   *)
END_FUNCTION_BLOCK

FUNCTION_BLOCK "DELAY_4"   // FB108, SCL
TITLE = DELAY_4
{ S7_Optimized_Access := 'FALSE' }
AUTHOR : hugo
FAMILY : SIGPRO
NAME : DELAY4
VERSION : 1.1
// this function block delays input values by each programm cycle
// after 4 cycles the in value has shifted to the out 4 and will be discarded after the next cycle
// the blocks can be cascaded.
   VAR_INPUT
      in : Real;
   END_VAR
   VAR_OUTPUT
      out1 : Real;
      out2 : Real;
      out3 : Real;
      out4 : Real;
   END_VAR
   VAR
      temp : Real;
   END_VAR
BEGIN


     #out4 := #out3;
     #out3 := #out2;
     #out2 := #out1;
     #out1 := #temp;
     #temp := #in;

   (* revision history

   hm 19.1.2007    rev 1.1
       added variable temp to add 1 delay  for q1

   *)
END_FUNCTION_BLOCK

FUNCTION_BLOCK "FADE"   // FB109, SCL
TITLE = FADE
{ S7_Optimized_Access := 'FALSE' }
AUTHOR : oscat
FAMILY : SIGPRO
NAME : FADE
VERSION : 1.3
// FADE is used to crossfade between the inputs IN1 and IN2. The fade_over time is specified with TF.
// When F = TRUE then Y = IN2 after the time TF, and when F = FALSE then Y = IN1.
// 
// uses: RMP_W [FB105]
//       _RMP_W [FB94] 
//       T_PLC_MS [FC64]
//       STIME [FB64],IDB_STIME [DB64]
   VAR_INPUT
      IN1 : Real;
      IN2 : Real;
      F : Bool;
      TF : Time;
      rst : Bool;
   END_VAR
   VAR_OUTPUT
      Y : Real;
   END_VAR
   VAR
      rmx : "RMP_W";
   END_VAR
BEGIN


   #rmx(RST := #rst AND NOT #F, SET := #rst AND #F, PT := #TF, UP := #F);
   #Y := (#IN2 - #IN1) / 65535.0 * DINT_TO_REAL(WORD_TO_DINT(#rmx.out)) + #IN1;


   (* code for rev 1.1
   IF rst THEN
       rmx(set := F, rst := NOT F);
   ELSIF F AND (NOT rmx.high) THEN
       rmx(PT := TF, UP := TRUE, e := TRUE, rst := FALSE, set := FALSE);
   ELSIF (NOT F) AND (NOT rmx.low) THEN
       rmx(PT := TF, UP := FALSE, e := TRUE, rst := FALSE, set := FALSE);
   ELSE
       rmx(e := FALSE, rst := FALSE, set := FALSE);
   END_IF;
   Y := (WORD_TO_REAL(rmx.out) * in1 + WORD_TO_REAL(FF - rmx.out) * IN2) / FF;
   *)


   (* revision history
   hm  26. dec 2007    rev 1.0
       original version

   hm  18. oct. 2008   rev 1.1
       improved performance
       changed calls for rmp_w because rmp_w has chaged

   hm  17. dec. 2008   rev 1.2
       function of input f was inverted

   hm  24. jan. 2009   rev 1.3
       delted unused var FF
   *)
END_FUNCTION_BLOCK

FUNCTION_BLOCK "FILTER_DW"   // FB110, SCL
TITLE = FILTER_DW
{ S7_Optimized_Access := 'FALSE' }
AUTHOR : hugo
FAMILY : SIGPRO
NAME : FILTDW
VERSION : 1.1
// FILTER_DW is an low pass filter with a programmable time T used for DWORD format.
// 
// uses: T_PLC_MS [FC64]
//       STIME [FB64],IDB_STIME [DB64]
   VAR_INPUT
      X : DWord;
      T : Time;
   END_VAR
   VAR_OUTPUT
      Y : DWord;
   END_VAR
   VAR
      last : DWord;
      tx : DWord;
      init : Bool;
      Yi : Real;
   END_VAR
   VAR_TEMP
      TOP_SI : Struct
         EV_CLASS : Byte;
         EV_NUM : Byte;
         PRIORITY : Byte;
         NUM : Byte;
         TYP2_3 : Byte;
         TYP1 : Byte;
         ZI1 : Word;
         ZI2_3 : DWord;
      END_STRUCT;
      START_UP_SI : Struct
         EV_CLASS : Byte;
         EV_NUM : Byte;
         PRIORITY : Byte;
         NUM : Byte;
         TYP2_3 : Byte;
         TYP1 : Byte;
         ZI1 : Word;
         ZI2_3 : DWord;
      END_STRUCT;
      ERR : Int;
   END_VAR
BEGIN


   (* read actual startup info *)
   (* OB1_SCAN_1  BYTE  -  B#16#01: Abschluss des Neustarts (Warmstarts)
                        -  B#16#02: Abschluss des Wiederanlaufs
                        -  B#16#03: Abschluss des freien Zyklus
                        -  B#16#04: Abschluss des Kaltstarts
                        -  B#16#05: Erster OB 1-Zyklus der neuen Master-CPU nach 
                                    Master-Reserve-Umschaltung und STOP des 
                                    bisherigen Masters *)

   #ERR := RD_SINFO (TOP_SI => #TOP_SI, START_UP_SI => #START_UP_SI);

   (* read system time *)
   #tx := "T_PLC_MS"();

   (* reset last_time on system startup *)
   IF #TOP_SI.EV_NUM = 1 OR #TOP_SI.EV_NUM = 2 OR #TOP_SI.EV_NUM = 4 THEN 
       #last := #tx;
   END_IF;

   (* startup initialisation *)
   IF NOT #init OR #T = t#0s THEN
       #init := TRUE;
       #Yi := DWORD_TO_REAL(#X);
   ELSE
       #Yi := #Yi + (DWORD_TO_REAL(#X) - DWORD_TO_REAL(#Y)) * DINT_TO_REAL(DWORD_TO_DINT(#tx) - DWORD_TO_DINT(#last)) / DINT_TO_REAL(T_CONV(#T));
   END_IF;
   #last := #tx;

   #Y := REAL_TO_DWORD(#Yi);


   (*
   hm 10. oct. 2008    rev 1.0
       original version

   hm  3. nov. 2008    REV 1.1
       corrected an overflow problem
   *)
END_FUNCTION_BLOCK

FUNCTION_BLOCK "FILTER_MAV_DW"   // FB111, SCL
TITLE = FILTER_MAV_DW
{ S7_Optimized_Access := 'FALSE' }
AUTHOR : hugo
FAMILY : SIGPRO
NAME : FIMAVDW
VERSION : 1.3
// FILTER_MAV_DW is a moving average filter with programmable length N for DWORD Data.
//  
// uses: INC1 [FC53]
   VAR_INPUT
      X : DWord;
      N : Int;
      RST : Bool;
   END_VAR
   VAR_OUTPUT
      Y : DWord;
   END_VAR
   VAR
      init : Bool;
      buffer : Array[0..31] of DWord;
      i : Int;
   END_VAR
   VAR_TEMP
      tmp : Int;
      tN : Int;
   END_VAR
BEGIN


   (* limit N to size of buffer *)
   #tN := MIN(IN1:=#N, IN2:=32);

   (* startup initialisation *)
   IF NOT #init OR #RST OR #tN = 0 THEN
       #init := TRUE;
       #tmp := #tN - 1;
       FOR #i := 0 TO #tmp DO
           #buffer[#i] := #X;
       END_FOR;
       #Y := #X;
   ELSE
       #tmp := #tN;
       #i := "INC1"(X:=#i, N:=#tmp);
       #Y := DINT_TO_DWORD(DWORD_TO_DINT(#Y) + (DWORD_TO_DINT(#X) - DWORD_TO_DINT(#buffer[#i])) / INT_TO_DINT(#tN));
       #buffer[#i] := #X;
   END_IF;


   (*
   hm 13. oct. 2008    rev 1.0
       original version

   hm  27. oct. 2008   rev 1.1
       added typecast to avoid warnings

   hm  24. nov. 2008   rev 1.2
       added typecasts to avoid warnings
       avoid divide by 0 if N = 0

   hm  23. feb. 2009   rev 1.3
       limit N to max array size

   *)
END_FUNCTION_BLOCK

FUNCTION_BLOCK "FILTER_MAV_W"   // FB112, SCL
TITLE = FILTER_MAV_W
{ S7_Optimized_Access := 'FALSE' }
AUTHOR : hugo
FAMILY : SIGPRO
NAME : FIMAVW
VERSION : 1.4
// FILTER_MAV_W is a moving average filter with programmable length N for WORD Data.
//  
// uses: INC1 [FC53]
   VAR_INPUT
      X : Word;
      N : Int;
      RST : Bool;
   END_VAR
   VAR_OUTPUT
      Y : Word;
   END_VAR
   VAR
      init : Bool;
      buffer : Array[0..31] of Word;
      i : Int;
      sum : DWord;
   END_VAR
   VAR_TEMP
      tmp : Int;
      tN : Int;
   END_VAR
BEGIN


   (* limit N to size of buffer *)
   #tN := MIN(IN1:=#N, IN2:=32);

   (* startup initialisation *)
   IF NOT #init OR #RST OR #tN = 0 THEN
     #init := TRUE;
     #tmp := #tN - 1;
     FOR #i := 0 TO #tmp DO
       #buffer[#i] := #X;
     END_FOR;
     #sum := DINT_TO_DWORD(WORD_TO_DINT(#Y) * INT_TO_DINT(#tN));
     #Y := #X;
   ELSE
     #tmp := #tN;
     #i := "INC1"(X:=#i, N:=#tmp);
     #sum := DINT_TO_DWORD(DWORD_TO_DINT(#sum) + WORD_TO_DINT(#X) - WORD_TO_DINT(#buffer[#i]));
     #Y := DINT_TO_WORD(DWORD_TO_DINT(#sum) / INT_TO_DINT(#tN));
     #buffer[#i] := #X;
   END_IF;


   (*
   hm 13. oct. 2008  rev 1.0
     original version

   hm  18. oct. 2008 rev 1.1
     added typecast to avoid warnings

   hm  24. nov. 2008 rev 1.2
     added typecasts to avoid warnings
     avoid devide by 0 if N = 0

   hm  23. feb. 2009 rev 1.3
     limit N to max array size

   hm  26. mar. 2011 rev 1.4
     corrected error in calculation
   *)
END_FUNCTION_BLOCK

FUNCTION_BLOCK "FILTER_W"   // FB113, SCL
TITLE = FILTER_W
{ S7_Optimized_Access := 'FALSE' }
AUTHOR : hugo
FAMILY : SIGPRO
NAME : FILTW
VERSION : 1.2
// FILTER_DW is an low pass filter with a programmable time T used for DWORD format.
// 
// uses: T_PLC_MS [FC64]
//       STIME [FB64],IDB_STIME [DB64]
   VAR_INPUT
      X : Word;
      T : Time;
   END_VAR
   VAR_OUTPUT
      Y : Word;
   END_VAR
   VAR
      last : DWord;
      tx : DWord;
      init : Bool;
      tmp : DWord;
   END_VAR
   VAR_TEMP
      TOP_SI : Struct
         EV_CLASS : Byte;
         EV_NUM : Byte;
         PRIORITY : Byte;
         NUM : Byte;
         TYP2_3 : Byte;
         TYP1 : Byte;
         ZI1 : Word;
         ZI2_3 : DWord;
      END_STRUCT;
      START_UP_SI : Struct
         EV_CLASS : Byte;
         EV_NUM : Byte;
         PRIORITY : Byte;
         NUM : Byte;
         TYP2_3 : Byte;
         TYP1 : Byte;
         ZI1 : Word;
         ZI2_3 : DWord;
      END_STRUCT;
      ERR : Int;
   END_VAR
BEGIN


   (* read actual startup info *)
   (* OB1_SCAN_1  BYTE  -  B#16#01: Abschluss des Neustarts (Warmstarts)
                        -  B#16#02: Abschluss des Wiederanlaufs
                        -  B#16#03: Abschluss des freien Zyklus
                        -  B#16#04: Abschluss des Kaltstarts
                        -  B#16#05: Erster OB 1-Zyklus der neuen Master-CPU nach 
                                    Master-Reserve-Umschaltung und STOP des 
                                    bisherigen Masters *)

   #ERR := RD_SINFO (TOP_SI => #TOP_SI, START_UP_SI => #START_UP_SI);

   (* read system time *)
   #tx := "T_PLC_MS"();

   (* reset last_time on system startup *)
   IF #TOP_SI.EV_NUM = 1 OR #TOP_SI.EV_NUM = 2 OR #TOP_SI.EV_NUM = 4 THEN 
     #init := false;
   END_IF;

   (* startup initialisation *)
   IF NOT #init OR #T = t#0s THEN
     #init := TRUE;
     #last := #tx;
     #Y := #X;
   ELSIF #Y = #X THEN
     #last := #tx;
   ELSE
     #tmp :=  DINT_TO_DWORD((WORD_TO_DINT(#X) - WORD_TO_DINT(#Y)) * (DWORD_TO_DINT(#tx) - DWORD_TO_DINT(#last)) / T_CONV(#T));
     IF #tmp <> 0 THEN
       #Y := DINT_TO_WORD(WORD_TO_DINT(#Y) + DWORD_TO_DINT(#tmp));
       #last := #tx;
     END_IF;
   END_IF;


   (*
   hm 10. oct. 2008  rev 1.0
     original version

   hm  3. nov. 2008  rev 1.1
     fixed overflow problem in formula

   hm  25. jan. 2011 rev 1.2
     fixed error in formula
   *)
END_FUNCTION_BLOCK

FUNCTION_BLOCK "FILTER_WAV"   // FB114, SCL
TITLE = FILTER_WAV
{ S7_Optimized_Access := 'FALSE' }
AUTHOR : hugo
FAMILY : SIGPRO
NAME : FILTWAV
VERSION : 1.2
// FILTER_WAV is a moving average filter with programmable length N for DWORD Data.
// 
// uses: INC1 [FC53]
//       DEC1 [FC52]
   VAR_INPUT
      X : Real;
      W : Array[0..15] of Real;
      RST : Bool;
   END_VAR
   VAR_OUTPUT
      Y : Real;
   END_VAR
   VAR
      init : Bool;
      buffer : Array[0..15] of Real;
      i : Int;
      n : Int;
   END_VAR
BEGIN


   (* startup initialisation *)
   IF NOT #init OR #RST THEN
       #init := TRUE;
       FOR #i := 0 TO 15 DO
           #buffer[#i] := #X;
       END_FOR;
       #i := 15;
       #Y := #X;
   ELSE
       #i := "INC1"(N:=16, X:=#i);
       #buffer[#i] := #X;
   END_IF;

   (* calculate the weighted average *)
   #Y := 0.0;
   FOR #n := 0 TO 15 DO
       #Y := #buffer[#i] * #W[#n] + #Y;
       #i := "DEC1"(N:=16, X:=#i);
   END_FOR;


   (*
   hm  14. oct. 2008   rev 1.0
       original version

   hm  27. oct. 2008   rev 1.1
       changed _DEC and _INC to DEC1 and INC1

   hm  10. mar. 2009   rev 1.2
       real constants updated to new systax using dot

   *)
END_FUNCTION_BLOCK

FUNCTION_BLOCK "SEL2_OF_3"   // FB115, SCL
TITLE = SEL2_OF_3
{ S7_Optimized_Access := 'FALSE' }
AUTHOR : oscat
FAMILY : SIGPRO
NAME : SEL2OF3
VERSION : 1.1
// SEL2_OF_3 checks if 3 input Signals are within a distance D from each other and calculates the average of the 3 inputs do not offset more than D from each other.
// If 1 input is more than D greater or smaller than any other input it will be ignored and the average will be calcualted from the remaining 2 Inputs.
// In the case the Output is only calculated from 2 Inputs a Warning Output W will display the Number of the discarded Input. if none of the 3 Inputs are within the allowed Delata D from each other, 
// an Error Output E is set True and the last valid Output will remain active until at least 2 Inputs are within a valid Range from each other.
   VAR_INPUT
      IN1 : Real;
      IN2 : Real;
      IN3 : Real;
      D : Real;
   END_VAR
   VAR_OUTPUT
      Y : Real;
      W : Int;
      "E" : Bool;
   END_VAR
   VAR
      D12 : Bool;
      D23 : Bool;
      D31 : Bool;
   END_VAR
BEGIN


   #D12 := ABS(#IN1-#IN2) <= #D;
   #D23 := ABS(#IN2-#IN3) <= #D;
   #D31 := ABS(#IN3-#IN1) <= #D;

   IF (#D12 AND #D23) OR (#D12 AND #D31) OR (#D23 AND #D31) THEN
       (* all 3 inputs are valid *)
       #Y := (#IN1 + #IN2 + #IN3) * 0.333333333333;
       #"E" := FALSE;
       #W := 0;
   ELSIF #D12 THEN
       (* only inut 1 and 2 are valid *)
       #Y := (#IN1 + #IN2) * 0.5;
       #"E" := FALSE;
       #W := 3;
   ELSIF #D23 THEN
       (* only inut 2 and 3 are valid *)
       #Y := (#IN2 + #IN3) * 0.5;
       #"E" := FALSE;
       #W := 1;
   ELSIF #D31 THEN
       (* only inut 3 and 1 are valid *)
       #Y := (#IN3 + #IN1) * 0.5;
       #"E" := FALSE;
       #W := 2;
   ELSE
       (* no calculation possible *)
       #"E" := TRUE;
       #W := 4;
   END_IF;


   (* revision history
   hm  18. may 2008    rev 1.0
       original version

   hm  10. mar. 2009   rev 1.1
       improved code
   *)
END_FUNCTION_BLOCK

FUNCTION_BLOCK "SEL2_OF_3B"   // FB116, SCL
TITLE = SEL2_OF_3B
{ S7_Optimized_Access := 'FALSE' }
AUTHOR : oscat
FAMILY : SIGPRO
NAME : SEL2OF3B
VERSION : 1.0
// SEL2_OF_3B is used to connect 3 binary sensors to one signal. the output Q reflects the state of at least two inputs.
// if two or more of the 3 inputs ate TRUE then Q will be TRUE and if two or more of the three inputs are FALSE then Q will be false.
// the main putrpose is the connection of 3 redundant binary sensors.  
// The output W will be active when one of the 3 inputs is of different state.
// to avoid flickering while the sensors are switching the output W will become active after a programmed delay of TD.
   VAR_INPUT
      IN1 : Bool;
      IN2 : Bool;
      IN3 : Bool;
      TD : Time;
   END_VAR
   VAR_OUTPUT
      Q : Bool;
      W : Bool;
   END_VAR
   VAR
      TDEL : TON;
   END_VAR
BEGIN


   #Q := (#IN1 AND #IN2) OR (#IN1 AND #IN3) OR (#IN2 AND #IN3);
   #TDEL(IN := (#IN1 XOR #IN2) OR (#IN1 XOR #IN3) OR (#IN2 XOR #IN3), PT := #TD);
   #W := #TDEL.Q;


   (* revision history
   hm      19. may 2008    rev 1.0
       original version

   *)
END_FUNCTION_BLOCK

FUNCTION_BLOCK "SH"   // FB117, SCL
TITLE = SH
{ S7_Optimized_Access := 'FALSE' }
AUTHOR : hugo
FAMILY : SIGPRO
NAME : SH
VERSION : 1.1
// this sample and hold module samples an input at the rising edge of clk an stores it in out.
// the out stays stable until the next rising clk edge appears.
// a trigger output as active for one cycle when the output was updated.
   VAR_INPUT
      in : Real;
      CLK : Bool;
   END_VAR
   VAR_OUTPUT
      out : Real;
      trig : Bool;
   END_VAR
   VAR
      edge : Bool;
   END_VAR
BEGIN


     IF #CLK AND NOT #edge THEN
         #out := #in;
         #trig := TRUE;
     ELSE;
         #trig := FALSE;
     END_IF;
     #edge := #CLK;

   (* revision history

   hm 16.1.2007    rev 1.1
       added trig output

   *)
END_FUNCTION_BLOCK

FUNCTION_BLOCK "SH_1"   // FB118, SCL
TITLE = SH_1
{ S7_Optimized_Access := 'FALSE' }
AUTHOR : hugo
FAMILY : SIGPRO
NAME : SH_1
VERSION : 1.2
// this sample and hold module samples an input every PT seconds.
// after a ample is taken the output Trig will be active for one cycle.
// 
// uses: T_PLC_MS [FC64]
//       STIME [FB64],IDB_STIME [DB64]
   VAR_INPUT
      in : Real;
      PT : Time;
   END_VAR
   VAR_OUTPUT
      out : Real;
      Trig : Bool;
   END_VAR
   VAR
      last : Time;
      tx : Time;
   END_VAR
   VAR_TEMP
      TOP_SI : Struct
         EV_CLASS : Byte;
         EV_NUM : Byte;
         PRIORITY : Byte;
         NUM : Byte;
         TYP2_3 : Byte;
         TYP1 : Byte;
         ZI1 : Word;
         ZI2_3 : DWord;
      END_STRUCT;
      START_UP_SI : Struct
         EV_CLASS : Byte;
         EV_NUM : Byte;
         PRIORITY : Byte;
         NUM : Byte;
         TYP2_3 : Byte;
         TYP1 : Byte;
         ZI1 : Word;
         ZI2_3 : DWord;
      END_STRUCT;
      ERR : Int;
   END_VAR
BEGIN


   (* OB1_SCAN_1  BYTE  -  B#16#01: Abschluss des Neustarts (Warmstarts)
                        -  B#16#02: Abschluss des Wiederanlaufs
                        -  B#16#03: Abschluss des freien Zyklus
                        -  B#16#04: Abschluss des Kaltstarts
                        -  B#16#05: Erster OB 1-Zyklus der neuen Master-CPU nach 
                                    Master-Reserve-Umschaltung und STOP des 
                                    bisherigen Masters *)

   #ERR := RD_SINFO (TOP_SI => #TOP_SI, START_UP_SI => #START_UP_SI);

   (* reset last_time on system startup *)
   IF #TOP_SI.EV_NUM = 1 OR #TOP_SI.EV_NUM = 2 OR #TOP_SI.EV_NUM = 4 THEN 
       #last := t#0ms;
   END_IF;

     (* read system time *)
     #tx := T_CONV(DWORD_TO_DINT("T_PLC_MS"()));

     IF #tx - #last >= #PT THEN
       #last := #tx;
       #out := #in;
       #Trig := TRUE;
     ELSE
       #Trig := FALSE;
     END_IF;

   (* revision history

   HM  6.1.2007  rev 1.1
     added trig output

   HM  17.9.2007  rev 1.2
     replaced time() with T_PLC_MS() for compatibility reasons
   *)
END_FUNCTION_BLOCK

FUNCTION_BLOCK "SH_2"   // FB119, SCL
TITLE = SH_2
{ S7_Optimized_Access := 'FALSE' }
AUTHOR : hugo
FAMILY : SIGPRO
NAME : SH_2
VERSION : 1.6
// this sample and hold module samples an input every PT seconds.
// this sample and hold also does avg and other calculations with the input data.
// an average is calculated while for this calculation disc samples are discarded,
// disc = 0 all samples are averaged,
// if disc = 1 the lowest value is ignored,
// if disc = 2 the lowest and highest values are ignored, 
// and so on.....
// 
// uses: T_PLC_MS [FC64]
//       STIME [FB64],IDB_STIME [DB64]
//       EVEN [FC76]
   VAR_INPUT
      in : Real;
      PT : Time;
      N : Int := 16;
      disc : Int;
   END_VAR
   VAR_OUTPUT
      out : Real;
      trig : Bool;
      avg : Real;
      high : Real;
      low : Real;
   END_VAR
   VAR
      "M" : Int;
      buf : Array[0..15] of Real;
      buf2 : Array[0..15] of Real;
      last : Time;
      i : Int;
      start : Int;
      temp : Real;
      stop : Int;
      tx : Time;
      d2 : Int;
   END_VAR
   VAR_TEMP
      TOP_SI : Struct
         EV_CLASS : Byte;
         EV_NUM : Byte;
         PRIORITY : Byte;
         NUM : Byte;
         TYP2_3 : Byte;
         TYP1 : Byte;
         ZI1 : Word;
         ZI2_3 : DWord;
      END_STRUCT;
      START_UP_SI : Struct
         EV_CLASS : Byte;
         EV_NUM : Byte;
         PRIORITY : Byte;
         NUM : Byte;
         TYP2_3 : Byte;
         TYP1 : Byte;
         ZI1 : Word;
         ZI2_3 : DWord;
      END_STRUCT;
      ERR : Int;
   END_VAR
BEGIN


   (* read actual startup info *)
   (* OB1_SCAN_1  BYTE  -  B#16#01: Abschluss des Neustarts (Warmstarts)
                        -  B#16#02: Abschluss des Wiederanlaufs
                        -  B#16#03: Abschluss des freien Zyklus
                        -  B#16#04: Abschluss des Kaltstarts
                        -  B#16#05: Erster OB 1-Zyklus der neuen Master-CPU nach 
                                    Master-Reserve-Umschaltung und STOP des 
                                    bisherigen Masters *)

   #ERR := RD_SINFO (TOP_SI => #TOP_SI, START_UP_SI => #START_UP_SI);

   (* reset last_time on system startup *)
   IF #TOP_SI.EV_NUM = 1 OR #TOP_SI.EV_NUM = 2 OR #TOP_SI.EV_NUM = 4 THEN 
       #last := t#0ms;
   END_IF;

   (* read system time *)
   #tx := T_CONV(DWORD_TO_DINT("T_PLC_MS"()));
   #d2 := WORD_TO_INT(SHR(IN:=INT_TO_WORD(#disc),N:=1));

   IF #tx - #last >= #PT THEN
       #last := #tx;
       #trig := TRUE;

       (* limit M to 0..16 *)
       #"M" := LIMIT(MN:=1,IN:=#N,MX:=16);

       (* edge detected lets take the sample *)
       FOR #i := #"M" - 1 TO 1 BY -1 DO #buf2[#i] := #buf2[#i-1]; END_FOR;
       #buf2[0] := #in;
       #out := #in;
       #buf BLKMOV #buf2;

       (* sort the ARRAY lowest value AT 0 *)
       FOR #start := 0 TO #"M" - 2 DO
         FOR #i := #start+1 TO #"M" - 1 DO
           IF #buf[#start] > #buf[#i] THEN
             #temp := #buf[#start];
             #buf[#start] := #buf[#i];
             #buf[#i] := #temp;
           END_IF;
         END_FOR;
       END_FOR;

       (* any calculation with the samples is here *)
       #stop := #"M" - 1 - #d2;
       #start := #d2;
       IF NOT "EVEN"(#disc) THEN #start := #start + 1; END_IF;
       #avg := 0;
       FOR #i := #start TO #stop DO #avg := #avg + #buf[#i]; END_FOR;
       #avg := #avg / INT_TO_REAL(#stop - #start +1);
       #low := #buf[#start];
       #high := #buf[#stop];
   ELSE
       #trig := FALSE;
   END_IF;


   (* revision history
   hm 20. jan. 2007    rev 1.1
       added input N to specify the amout of samples for average and high low calculations
       added trig output

   hm 10. sep. 2007    rev 1.2
       an error would be generated if N was set to 0, now n is forced to1 if set to 0.
       index was out of array.

   hm  17. sep. 2007   rev 1.3
       replaced time() with t_plc_ms() for compatibility reasons

   hm  6. jan. 2008    rev 1.4
       improved performance

   hm  14. jun. 2008   rev 1.5
       set default for input N = 16

   hm  10. mar. 2009   rev 1.6
       added type conversion for compatibility reasons

   *)
END_FUNCTION_BLOCK

FUNCTION_BLOCK "SH_T"   // FB120, SCL
TITLE = SH_T
{ S7_Optimized_Access := 'FALSE' }
AUTHOR : hugo
FAMILY : SIGPRO
NAME : SH_T
VERSION : 1.1
// this sample and hold module samples an input while en is high.
// during the high time of en the output follows in.
// the out stays stable until the en goes high again.
   VAR_INPUT
      IN : Real;
      "E" : Bool;
   END_VAR
   VAR_OUTPUT
      OUT : Real;
   END_VAR
BEGIN


   IF #"E" THEN #OUT := #IN; END_IF;

   (* revision history
   hm  1. sep. 2006    rev 1.0
       original version

   hm  18. oct. 2008   rev 1.1
       changed input en to e for compatibility reasons

   *)
END_FUNCTION_BLOCK

FUNCTION_BLOCK "STAIR2"   // FB121, SCL
TITLE = STAIR2
{ S7_Optimized_Access := 'FALSE' }
AUTHOR : oscat
FAMILY : SIGPRO
NAME : STAIR2
VERSION : 1.4
// the function stair2 converts an anlog input signal to a staircase like output.
// D is the step width for the output signal. the output will use D as a hysteresis for a stairchange.
// if D = 0 then the output follows the input without a chage.
// 
// uses: FLOOR [FC81]
   VAR_INPUT
      X : Real;
      D : Real;
   END_VAR
   VAR_OUTPUT
      Y : Real;
   END_VAR
BEGIN


   IF #D > 0.0 THEN
       IF #X >= #Y + #D OR #X <= #Y - #D THEN #Y := "FLOOR"(#X/#D) * #D; END_IF;
   ELSE
       #Y := #X;
   END_IF;


   (* revision history
   hm  28 jan 2007     rev 1.0
       original version

   hm  27. dec 2007    rev 1.1
       changed code for better performance

   hm  30. jun. 2008   rev 1.2
       added type conversions to avoid warnings under codesys 3.0

   ks  26. oct. 2008   rev 1.3
       improved code

   hm  10. mar. 2009   rev 1.4
       real constants updated to new systax using dot

   *)
END_FUNCTION_BLOCK

FUNCTION_BLOCK "FILTER_I"   // FB238, SCL
TITLE = FILTER_I
{ S7_Optimized_Access := 'FALSE' }
AUTHOR : hugo
FAMILY : SIGPRO
NAME : FILTI
VERSION : 1.0
// FILTER_I is a low pass filter with a programmable time T used for INT format.
//  
// uses: T_PLC_MS [FC64]
//       STIME [FB64],IDB_STIME [DB64]
   VAR_INPUT
      X : Int;
      T : Time;
   END_VAR
   VAR_OUTPUT
      Y : Int;
   END_VAR
   VAR
      Yi : DInt;
      last : DWord;
      tx : DWord;
      init : Bool;
   END_VAR
   VAR_TEMP
      TOP_SI : Struct
         EV_CLASS : Byte;
         EV_NUM : Byte;
         PRIORITY : Byte;
         NUM : Byte;
         TYP2_3 : Byte;
         TYP1 : Byte;
         ZI1 : Word;
         ZI2_3 : DWord;
      END_STRUCT;
      START_UP_SI : Struct
         EV_CLASS : Byte;
         EV_NUM : Byte;
         PRIORITY : Byte;
         NUM : Byte;
         TYP2_3 : Byte;
         TYP1 : Byte;
         ZI1 : Word;
         ZI2_3 : DWord;
      END_STRUCT;
      ERR : Int;
   END_VAR
BEGIN


   (* read actual startup info *)
   (* OB1_SCAN_1  BYTE  -  B#16#01: Abschluss des Neustarts (Warmstarts)
                        -  B#16#02: Abschluss des Wiederanlaufs
                        -  B#16#03: Abschluss des freien Zyklus
                        -  B#16#04: Abschluss des Kaltstarts
                        -  B#16#05: Erster OB 1-Zyklus der neuen Master-CPU nach 
                                    Master-Reserve-Umschaltung und STOP des 
                                    bisherigen Masters *)

   #ERR := RD_SINFO (TOP_SI => #TOP_SI, START_UP_SI => #START_UP_SI);

   (* read system time *)
   #tx := "T_PLC_MS"();

   (* reset last_time on system startup *)
   IF #TOP_SI.EV_NUM = 1 OR #TOP_SI.EV_NUM = 2 OR #TOP_SI.EV_NUM = 4 THEN 
       #last := #tx;
   END_IF;

   (* startup initialisation *)
   IF NOT #init OR #T = t#0s THEN
       #init := TRUE;
       #Yi := INT_TO_DINT(#X) * 1000;
   ELSE
       (* to increase accuracy of the filter we calculate internal Yi wich is Y * 1000 *)
       #Yi := #Yi + INT_TO_DINT(#X - #Y) * (DWORD_TO_DINT(#tx) - DWORD_TO_DINT(#last)) * 1000 / T_CONV(#T);
   END_IF;
   #last := #tx;
   #Y := DINT_TO_INT(#Yi / 1000);


   (*
   hm 8. nov. 2008 rev 1.0
       original version

   *)
END_FUNCTION_BLOCK

FUNCTION_BLOCK "TREND_DW"   // FB245, SCL
TITLE = TREND_DW
{ S7_Optimized_Access := 'FALSE' }
AUTHOR : hugo
FAMILY : SIGPRO
NAME : TREND_DW
VERSION : 1.2
// trend_DW analyses the trend of a input signal.
// The Output Q is True if the input X is >= last_X and is false if the input X is <= last_X
// in addition to the trend the output TU will be high for one cycle to signal a rising of the input value X
// and  TD will signal a decreasing value on the input X.
// in case of a change the output D will show the delta of the input to the last input value.
   VAR_INPUT
      X : DWord;
   END_VAR
   VAR_OUTPUT
      Q : Bool;
      TU : Bool;
      TD : Bool;
      D : DWord;
   END_VAR
   VAR
      last_X : DWord;
   END_VAR
BEGIN


   IF DWORD_TO_DINT(#X) > DWORD_TO_DINT(#last_X) THEN
       #TU := TRUE;
       #TD := FALSE;
       #D := DINT_TO_DWORD(DWORD_TO_DINT(#X) - DWORD_TO_DINT(#last_X));
       #Q := TRUE;
   ELSIF DWORD_TO_DINT(#X) < DWORD_TO_DINT(#last_X) THEN
       #TD := TRUE;
       #TU := FALSE;
       #D := DINT_TO_DWORD(DWORD_TO_DINT(#last_X) - DWORD_TO_DINT(#X));
       #Q := FALSE;
   ELSE
       #TU := FALSE; 
       #TD := FALSE;
       #D := 0;
   END_IF;
   #last_X := #X;


   (* revision history
   hm  21. nov. 2008   rev 1.0
       original version

   hm  20. feb. 2009   rev 1.1
       added outputs TU, TD and D

   hm  14. mar. 2009   rev 1.2
       removed double assignments

   *)
END_FUNCTION_BLOCK

FUNCTION_BLOCK "TREND"   // FB251, SCL
TITLE = TREND
{ S7_Optimized_Access := 'FALSE' }
AUTHOR : hugo
FAMILY : SIGPRO
NAME : TREND
VERSION : 1.0
// trend analyses the trend of a input signal.
// The Output Q is True if the input X is >= last_X and is false if the input X is <= last_X
// in addition to the trend the output TU will be high for one cycle to signal a rising of the input value X
// and  TD will signal a decreasing value on the input X.
// in case of a change the output D will show the delta of the input to the last input value.
   VAR_INPUT
      X : Real;
   END_VAR
   VAR_OUTPUT
      Q : Bool;
      TU : Bool;
      TD : Bool;
      D : Real;
   END_VAR
   VAR
      last_X : Real;
   END_VAR
BEGIN


   #TU := #X > #last_X;
   #TD := #X < #last_X;
   #Q := #TU OR #TD;
   #D := #X - #last_X;

   #last_X := #X;



   (* revision history
   hm 21. aug. 2009 rev 1.0
    original version

   *)
END_FUNCTION_BLOCK

FUNCTION "DEC1" : Int   // FC52, SCL
TITLE = DEC1
{ S7_Optimized_Access := 'FALSE' }
AUTHOR : hugo
FAMILY : MATH
NAME : DEC1
VERSION : 1.1
// This is a decrement function which decrements the variable X by 1 and if 0 is reached, it begins with M again.
// _dec1(3,X) will generate 3,2,1,0,3,2,...
   VAR_INPUT
      X : Int;
      N : Int;
   END_VAR
BEGIN


   IF #X = 0 THEN
       #DEC1 := #N - 1;
   ELSE
       #DEC1 := #X - 1;
   END_IF;

   (* this is a very elegant version but 50% slower
   X := (X - 1 + N) MOD N;
   *)


   (* revision history
   hm  13. oct. 2008   rev 1.0
       original version

   hm  27. oct. 2008   rev 1.1
       added statement to return value for compatibility reasons
   *)
END_FUNCTION

FUNCTION "INC1" : Int   // FC53, SCL
TITLE = INC1
{ S7_Optimized_Access := 'FALSE' }
AUTHOR : hugo
FAMILY : MATH
NAME : INC1
VERSION : 1.2
// This is a increment function which increments the variable X by 1 and if M is reached, it begins with 0 again.
// _inc1(3,X) will generate 0,1,2,3,0,1,.....
   VAR_INPUT
      X : Int;
      N : Int;
   END_VAR
BEGIN


   IF #X >= #N - 1 THEN
       #INC1 := 0;
   ELSE
       #INC1 := #X + 1;
   END_IF;


   (* this elegant version is 50% slower
   INC1 := X := (x + 1) MOD N;
   *)



   (* revision history
   hm  13. oct. 2008   rev 1.0
       original version

   hm  22. oct. 2008   rev 1.1
       added statement to return value for compatibility reasons

   hm  23. feb. 2009   rev 1.2
       when inc1 is called with X >= N inc will continue with 0
   *)
END_FUNCTION

FUNCTION "T_PLC_MS" : DWord   // FC64, SCL
TITLE = T_PLC_MS
{ S7_Optimized_Access := 'FALSE' }
AUTHOR : hugo
FAMILY : MEASURE
NAME : T_PLC_MS
VERSION : 1.2
// T_PLC_MS reads the internal PLC timer and return the time, it has the advantage to be able to set a debug mode 
// and speed up the counter to test the plc timer overrun which occurs every 50 days respectively 25 days at siemens S7
// this routine also allows to correct the behavior of s7 where the internal plc counter will not count all 32 bits.
// 
// uses: STIME [FB64],IDB_STIME [DB64]
BEGIN


   "IDB_STIME"(); 
   #T_PLC_MS := "IDB_STIME".tx; 
   (* hier muss die korrektur für step7 stattfinden
   plctime muss den vollen wertebereich von time ausnutzen:
   wenn bei step7 time -24tage bis plus 24 tage ist dann muss der timer auch beim überlauf auf -24tage springen 
   und auf keinen fall auf 0 !!!!
   für siemens muss ein weiterer fb im main eingebunden werden der sicherstellt das alle 32 bits durchgezählt werden.
   es kann nur ein fb sein den er muss sich das oberste (32te) bit merken.
   oder etwa spring s7 bei überlauf auf -24 tage????? dann wäre keine korrektur nötig.
   *)
   IF "debug" THEN
       #T_PLC_MS := DINT_TO_DWORD((DWORD_TO_DINT(SHL(IN:=#T_PLC_MS,N:="N") OR SHL(IN:=DWORD#1,N:="N"))-1) + DWORD_TO_DINT("offset_FC64_1"));
   END_IF;


   (* revision history
   hm  14.9.2007   rev 1.0
       original version

   hm  12. nov 2007    rev 1.1
       added temporaray variable tx because some compilers could not handle time() as an argument

   hm  16. nov. 2008   rev 1.2
       initialized constants with 0 for compatibility reasons
   *)
END_FUNCTION

FUNCTION "EVEN" : Bool   // FC76, SCL
TITLE = EVEN
{ S7_Optimized_Access := 'FALSE' }
AUTHOR : hugo
FAMILY : MATH
NAME : EVEN
VERSION : 1.2
// this function chacks an input for even value
// the output is true if the input is even.
   VAR_INPUT
      in : DInt;
   END_VAR
   VAR_TEMP
      tIN : DInt;
      _IN AT tIN : Array[0..31] of Bool;
   END_VAR
BEGIN


   #tIN := #in;
   #EVEN := NOT #_IN[24]; //EVEN := NOT in.0;

   (* revision history
   hm  1. oct 2006 rev 1.0
     ORIGINAL VERSION

   hm  01.12.2007  rev 1.1
     changed code for improved performance

   hm  21. mar. 2008 rev 1.2
     changed type of input IN from INT to DINT
   *)
END_FUNCTION

FUNCTION "FLOOR" : Int   // FC81, SCL
TITLE = FLOOR
{ S7_Optimized_Access := 'FALSE' }
AUTHOR : hugo
FAMILY : MATH
NAME : FLOOR
VERSION : 1.1
// This is a rounding function which returns the biggest possible integer which is less or equal to X.
// floor(3.14) = 3
// floor(-3.14) = 4
   VAR_INPUT
      X : Real;
   END_VAR
BEGIN


   #FLOOR := REAL_TO_INT(#X);
   IF #FLOOR > #X THEN
       #FLOOR := #FLOOR - 1;
   END_IF;

   (* revision history
   hm    7. feb 2007   rev 1.0
     originlal version

   hm    21. mar. 2008 rev 1.1
     replaced trunc with real_to_int for compatibility reasons

   *)
END_FUNCTION

FUNCTION "SIGN_R" : Bool   // FC109, SCL
TITLE = SIGN_R
{ S7_Optimized_Access := 'FALSE' }
AUTHOR : hugo
FAMILY : MATH
NAME : SIGN_R
VERSION : 1.4
// this function return true if the real input is negative
   VAR_INPUT
      in : Real;
   END_VAR
BEGIN


   #SIGN_R := #in < 0.0;


   (* revision history
   hm 19.1.2007    rev 1.1
       changed method of function for better compatibility to other systems

   hm  1.12.2007   rev 1.2
       changed code to improve performance

   hm  14. jun. 2008   rev 1.3
       improved performace

   hm 10. mar. 2009    rev 1.4
       real constants updated to new systax using dot
   *)
END_FUNCTION

FUNCTION "AIN" : Real   // FC317, SCL
TITLE = AIN
{ S7_Optimized_Access := 'FALSE' }
AUTHOR : oscat
FAMILY : SIGPRO
NAME : AIN
VERSION : 1.5
// Ain converts signals from A/D converters or other analog sources to an internal real value
// the lowest number of bits are extracted from the input word and the sign will be extracted if available separately.
// the output signal is then conditioned to range from low to high values for a 0 to max value on the analog inputs:
// for example a 15bit input (bits := 12) with sign at bit 15 (0..15) will deliver 0.0 (low value at 0) for an input value of 2#0000_0000_0000
// an input value of 2#1111_1111_1111 will deliver 10.0 on the output (high value set to 10).
   VAR_INPUT
      in : DWord;
      Bits : Byte;
      sign : Byte;
      low : Real;
      high : Real;
   END_VAR
   VAR_TEMP
      temp1 : DWord;
      ttemp1 AT temp1 : Array[0..31] of Bool;
      temp2 : DWord;
      sx : Bool;
   END_VAR
BEGIN


     (* extract the sign bit *)
     IF BYTE_TO_INT(#sign) < 32 THEN
         #temp1 := SHR(IN:=#in,N:=BYTE_TO_INT(#sign));
         #sx := #ttemp1[24];
     ELSE
         #sx := FALSE;
     END_IF;
     #temp1 := SHR(IN:="ff",N:=32-BYTE_TO_INT(#Bits));
     #temp2 := #in AND #temp1;
     #AIN := (#high - #low) * DWORD_TO_REAL(#temp2) / DWORD_TO_REAL(#temp1) + #low;
     IF #sx THEN #AIN := -#AIN; END_IF;

   (* revision history
   hm 18.8.2006    rev 1.1
       fixed an error with low value negative and high value 0.

   hm 19.1.2007    rev 1.2
       fixed an error with sign bit.

   hm  13.9.2007   rev 1.3
       changed code to avoid warning under codesys 2.8.1

   hm  2. dec 2007 rev 1.4
       changed code for better performance

   hm  16. mar 2008    rev 1.5
       added type conversions to avoid warnings under codesys 30
   *)
END_FUNCTION

FUNCTION "AOUT" : DWord   // FC318, SCL
TITLE = AOUT
{ S7_Optimized_Access := 'FALSE' }
AUTHOR : oscat
FAMILY : SIGPRO
NAME : AOUT
VERSION : 1.4
// this module conditions an internal real value for a signal output D/A converter.
// Aout converts and internal real value to a word for an D/A converter or other output devices.
// The input value is converted to a n-bit wide output and a sign bit is set separately as specified.
// the outout min value is set for the specified min input value and the max output is set for the max input value.
// an input higher or lower then the max or min value will set the respective max or min value or the output.
// 
// uses: SIGN_R [FC109]
   VAR_INPUT
      in : Real;
      Bits : Byte;
      sign : Byte;
      low : Real;
      high : Real;
   END_VAR
   VAR_TEMP
      in2 : Real;
      sx : Bool;
   END_VAR
BEGIN


     (* if sign bit is defined *)
     IF WORD_TO_INT(BYTE_TO_WORD(#sign)) < 32 THEN
         #sx := "SIGN_R"(in:=#in);
         #in2 := ABS(#in);
     ELSE
         #in2 := #in;
     END_IF;

     (* begrenze in auf die zulässigen werte *)
     #in2 := LIMIT(MN:=#low,IN:=#in2,MX:=#high);

     (* Berechne den Ausgnagswert *)
     #AOUT := DINT_TO_DWORD(REAL_TO_DINT((#in2 - #low) / (#high - #low) * (DINT_TO_REAL(DWORD_TO_DINT(SHL(IN:="ff_FC318",N:=BYTE_TO_INT(#Bits)))) -1)));
     IF #sx THEN #AOUT := SHL(IN:="ff_FC318",N:=WORD_TO_INT(BYTE_TO_WORD(#sign))) OR #AOUT; END_IF;

   (*
   revision history

   hm 18.1.2007    rev 1.1
     renamed Modul to aout.
     changed Output to 32 Bit max.
     corrected error with sign bit.

   hm  13.9.2007   rev 1.2
     changed code to avoid warning under codesys 2.8.1

   hm  2. dec 2007   rev 1.3
     changed code for better performance

   hm  23. feb 2008  rev 1.4
     changed code for better performance
   *)
END_FUNCTION

FUNCTION "BYTE_TO_RANGE" : Real   // FC320, SCL
TITLE = BYTE_TO_RANGE
{ S7_Optimized_Access := 'FALSE' }
AUTHOR : hugo
FAMILY : SIGPRO
NAME : BY2RA
VERSION : 1.0
// Byte_to_Range converts a Byte into a real between low and high.
   VAR_INPUT
      X : Byte;
      low : Real;
      high : Real;
   END_VAR
BEGIN


     #BYTE_TO_RANGE := (#high - #low) * DINT_TO_REAL(BYTE_TO_DINT(#X)) / 255.0 + #low;


   (* revision history
   hm  9. jan 2008   rev 1.0
     original version

   *)
END_FUNCTION

FUNCTION "MIX" : Real   // FC321, SCL
TITLE = MIX
{ S7_Optimized_Access := 'FALSE' }
AUTHOR : hugo
FAMILY : SIGPRO
NAME : MIX
VERSION : 1.1
// MIX is an analog Mixer. The Output is (1-M)*A + M*B.
   VAR_INPUT
      "A" : Real;
      "B" : Real;
      "M" : Real;
   END_VAR
BEGIN


   #MIX := (1.0 - #"M") * #"A" + #"M" * #"B";


   (* revision history
   hm  19. Nov 2007    rev 1.0
       original version

   hm  10. mar 2009    rev 1.1
       real constants updated to new systax using dot

   *)
END_FUNCTION

FUNCTION "MUX_R2" : Real   // FC322, SCL
TITLE = MUX_R2
{ S7_Optimized_Access := 'FALSE' }
AUTHOR : oscat
FAMILY : SIGPRO
NAME : MUX_R2
VERSION : 1.1
// MUX_R2 is an analog Multiplexer.
// one of 2 real inputs are selected and put through to out.
// The Adress input A selects between 2 Real inputs IN0 and IN1, A=0 > In0, A=1 > in1.
   VAR_INPUT
      IN0 : Real;
      IN1 : Real;
      "A" : Bool;
   END_VAR
BEGIN


   #MUX_R2 := SEL(G:=#"A", IN0:=#IN0, IN1:=#IN1);


   (* revision history
   hm  19. jan. 2007   rev 1.0
       original version

   hm  16. oct. 2008   rev 1.1
       improved performance


   *)
END_FUNCTION

FUNCTION "MUX_R4" : Real   // FC323, SCL
TITLE = MUX_R4
{ S7_Optimized_Access := 'FALSE' }
AUTHOR : oscat
FAMILY : SIGPRO
NAME : MUX_R4
VERSION : 1.1
// MUX_R4 is an analog Multiplexer.
// one of 4 real inputs are selected and put through to out.
// The Adress input A0 and A1 selects between the 4 Real inputs IN0.. IN1.
   VAR_INPUT
      IN0 : Real;
      IN1 : Real;
      IN2 : Real;
      IN3 : Real;
      A0 : Bool;
      A1 : Bool;
   END_VAR
BEGIN


   IF #A1 THEN
       #MUX_R4 := SEL(G:=#A0, IN0:=#IN2, IN1:=#IN3);
   ELSE
       #MUX_R4 := SEL(G:=#A0, IN0:=#IN0, IN1:=#IN1);
   END_IF;



   (* revision history
   hm  19. jan 2007    rev 1.0
       original version

   hm  16. oct. 2008   rev 1.1
       improved performance
   *)
END_FUNCTION

FUNCTION "OFFSET" : Real   // FC324, SCL
TITLE = OFFSET
{ S7_Optimized_Access := 'FALSE' }
AUTHOR : oscat
FAMILY : SIGPRO
NAME : OFFSET
VERSION : 1.0
// The Function offset adds offsets to an analog signal depending on digital inputs.
// all selected offsets are added at the same time.
// with the input D a default value instead of the input X can be used.
   VAR_INPUT
      X : Real;
      O1 : Bool;
      O2 : Bool;
      O3 : Bool;
      O4 : Bool;
      D : Bool;
      Offset_1 : Real;
      Offset_2 : Real;
      Offset_3 : Real;
      Offset_4 : Real;
      default : Real;
   END_VAR
BEGIN


   IF #D THEN #OFFSET := #default; ELSE #OFFSET := #X; END_IF;
   IF #O1 THEN #OFFSET := #OFFSET + #Offset_1; END_IF;
   IF #O2 THEN #OFFSET := #OFFSET + #Offset_2; END_IF;
   IF #O3 THEN #OFFSET := #OFFSET + #Offset_3; END_IF;
   IF #O4 THEN #OFFSET := #OFFSET + #Offset_4; END_IF;
END_FUNCTION

FUNCTION "OFFSET2" : Real   // FC325, SCL
TITLE = OFFSET2
{ S7_Optimized_Access := 'FALSE' }
AUTHOR : oscat
FAMILY : SIGPRO
NAME : OFFSET2
VERSION : 1.0
// The Function offset adds offsets to an analog signal depending on digital inputs.
// one offset can be added at the same time, if more then one input is true, the one with the highest number (o1 .. o4) will be used.
// The input D will select a default value instead of X for input.
   VAR_INPUT
      X : Real;
      O1 : Bool;
      O2 : Bool;
      O3 : Bool;
      O4 : Bool;
      D : Bool;
      Offset_1 : Real;
      Offset_2 : Real;
      Offset_3 : Real;
      Offset_4 : Real;
      default : Real;
   END_VAR
BEGIN


     IF #D THEN #OFFSET2 := #default; ELSE #OFFSET2 := #X; END_IF;
     IF #O4 THEN #OFFSET2 := #OFFSET2 + #Offset_4;
     ELSIF #O3 THEN #OFFSET2 := #OFFSET2 + #Offset_3;
     ELSIF #O2 THEN #OFFSET2 := #OFFSET2 + #Offset_2;
     ELSIF #O1 THEN #OFFSET2 := #OFFSET2 + #Offset_1;
     END_IF;
END_FUNCTION

FUNCTION "OVERRIDE" : Real   // FC326, SCL
TITLE = OVERRIDE
{ S7_Optimized_Access := 'FALSE' }
AUTHOR : oscat
FAMILY : SIGPRO
NAME : OVERRIDE
VERSION : 1.0
// OVERRIDE deliveres the maximum absolute value of the 3 inputs X1, X2 and X3.
// with the inputs E1, E2 and E3 each of the 3 inputs can be turned on or off.
   VAR_INPUT
      X1 : Real;
      X2 : Real;
      X3 : Real;
      E1 : Bool;
      E2 : Bool;
      E3 : Bool;
   END_VAR
BEGIN


   IF #E1 THEN #OVERRIDE := #X1; END_IF;
   IF #E2 AND ABS(#X2) > ABS(#OVERRIDE) THEN #OVERRIDE := #X2; END_IF;
   IF #E3 AND ABS(#X3) > ABS(#OVERRIDE) THEN #OVERRIDE := #X3; END_IF;

   (* revision history
   hm    4.11.2007        rev 1.0
       original version

   *)
END_FUNCTION

FUNCTION "RANGE_TO_BYTE" : Byte   // FC327, SCL
TITLE = RANGE_TO_BYTE
{ S7_Optimized_Access := 'FALSE' }
AUTHOR : hugo
FAMILY : SIGPRO
NAME : RA2BY
VERSION : 1.0
// Range_to_byte converts a real value between low and high into a byte
   VAR_INPUT
      X : Real;
      low : Real;
      high : Real;
   END_VAR
BEGIN


     #RANGE_TO_BYTE := INT_TO_BYTE(REAL_TO_INT(DINT_TO_REAL(TRUNC((LIMIT(MN:=#low,IN:=#X,MX:=#high)-#low))) * 255.0 / (#high - #low)));


   (* revision history
   hm  9. jan 2008   rev 1.0
     original version

   *)
END_FUNCTION

FUNCTION "RANGE_TO_WORD" : Word   // FC328, SCL
TITLE = RANGE_TO_WORD
{ S7_Optimized_Access := 'FALSE' }
AUTHOR : hugo
FAMILY : SIGPRO
NAME : RA2WO
VERSION : 1.0
// Range_to_word converts a real value between low and high into a byte
   VAR_INPUT
      X : Real;
      low : Real;
      high : Real;
   END_VAR
BEGIN


     #RANGE_TO_WORD := DINT_TO_WORD(REAL_TO_DINT(DINT_TO_REAL(TRUNC((LIMIT(MN:=#low,IN:=#X,MX:=#high)-#low))) * 65535.0 / (#high - #low)));


   (* revision history
   hm  9. jan 2008   rev 1.0
     original version

   *)
END_FUNCTION

FUNCTION "SCALE" : Real   // FC329, SCL
TITLE = SCALE
{ S7_Optimized_Access := 'FALSE' }
AUTHOR : hugo
FAMILY : SIGPRO
NAME : SCALE
VERSION : 1.0
// Scale is used to translate an input x to output by the formula Y = X*K + O.
// at the same time the output is limited to MN and MX.
   VAR_INPUT
      X : Real;
      K : Real;
      O : Real;
      MX : Real;
      MN : Real;
   END_VAR
BEGIN


   #SCALE := LIMIT(MN:=#MN,IN:=#X * #K + #O,MX:=#MX);


   (* revision history
   hm  16. may. 2008       rev 1.0
       original version
   *)
END_FUNCTION

FUNCTION "SCALE_B" : Real   // FC330, SCL
TITLE = SCALE_B
{ S7_Optimized_Access := 'FALSE' }
AUTHOR : hugo
FAMILY : SIGPRO
NAME : SCALEB
VERSION : 1.1
// Scale_B is used to translate and scale a byte input x to a real output.
   VAR_INPUT
      X : Byte;
      I_LO : Byte;
      I_HI : Byte;
      O_LO : Real;
      O_HI : Real;
   END_VAR
BEGIN


     IF #I_HI = #I_LO THEN
       #SCALE_B := #O_LO;
     ELSE
       #SCALE_B := (#O_HI - #O_LO) / (BYTE_TO_INT(#I_HI) - BYTE_TO_INT(#I_LO)) * LIMIT(MN:=BYTE_TO_INT(#I_LO),IN:=BYTE_TO_INT(#X),MX:=BYTE_TO_INT(#I_HI));
     END_IF;


   (* revision history
   hm  18. may. 2008   rev 1.0
     original version

   hm  18. jan 2011    rev 1.1
     avoid division by 0

   *)
END_FUNCTION

FUNCTION "SCALE_B2" : Real   // FC331, SCL
TITLE = SCALE_B2
{ S7_Optimized_Access := 'FALSE' }
AUTHOR : hugo
FAMILY : SIGPRO
NAME : SCALEB2
VERSION : 1.4
// version 1.4 3. nov. 2008
// programmer  hugo
// tested by   dalbi
// 
// this functiob block can scale up to two inputs.
// the inputs have their min value at 0 and their max value at 255 while the min and max value can be either positive or negative.
// the inputs ramp between min and max values for the respective inputs to be between (0..255).
// the summed output is then scaled by an scale input K and a offset O can be added to the output.
// the min and max input configurations can be edited in the cfc editor by double clicking the symbol body.
   VAR_INPUT
      in1 : Byte;
      in2 : Byte;
      K : Real;
      O : Real;
      in1_min : Real;
      in1_max : Real;
      in2_min : Real;
      in2_max : Real;
   END_VAR
BEGIN


   #SCALE_B2 := (((#in1_max - #in1_min)* INT_TO_REAL(BYTE_TO_INT(#in1)) + 
               (#in2_max - #in2_min)* INT_TO_REAL(BYTE_TO_INT(#in2))) * 
               0.003921569 + #in1_min + #in2_min) * #K + #O;


   (* code bofore rev 1.2
   scale_B2 :=     ((in1_max - in1_min)* in1 / 255 + in1_min +
                   (in2_max - in2_min)* in2 / 255 + in2_min)
                   * K + O;
   *)

   (* revision History
   hm 19.1.2007        rev 1.1
       changed outputs to real to avoid overflow of integer
       added offset for better cascading of scale functions
       changed from FB to function

   hm  6. jan 2008     rev 1.2
       improved performance

   hm  26. oct. 2008   rev 1.3
       code optimization

   hm  3. nov. 2008    rev 1.4
       used wrong factor in formula

   *)
END_FUNCTION

FUNCTION "SCALE_B4" : Real   // FC332, SCL
TITLE = SCALE_B4
{ S7_Optimized_Access := 'FALSE' }
AUTHOR : hugo
FAMILY : SIGPRO
NAME : SCALEB4
VERSION : 1.4
// this functiob block can scale up to 4 inputs.
// the inputs have their min value at 0 and their max value at 255 while the min and max value can be either positive or negative.
// the inputs ramp between min and max values for the respective inputs to be between (0..255).
// the summed output is then scaled by an scale input K and a offset O can be added to the output.
// the min and max input configurations can be edited in the cfc editor by double clicking the symbol body.
   VAR_INPUT
      in1 : Byte;
      in2 : Byte;
      in3 : Byte;
      in4 : Byte;
      K : Real;
      O : Real;
      in1_min : Real;
      in1_max : Real;
      in2_min : Real;
      in2_max : Real;
      in3_min : Real;
      in3_max : Real;
      in4_min : Real;
      in4_max : Real;
   END_VAR
BEGIN


   #SCALE_B4 := (((#in1_max - #in1_min)* INT_TO_REAL(BYTE_TO_INT(#in1)) + 
               (#in2_max - #in2_min)* INT_TO_REAL(BYTE_TO_INT(#in2)) + 
               (#in3_max - #in3_min)* INT_TO_REAL(BYTE_TO_INT(#in3)) + 
               (#in4_max - #in4_min)* INT_TO_REAL(BYTE_TO_INT(#in4)))* 
               0.003921569 + #in1_min + #in2_min + #in3_min + #in4_min) * #K + #O;


   (* revision History
   hm 19.1.2007        rev 1.1
       changed outputs to real to avoid overflow of integer
       added offset for better cascading of scale functions
       changed from fb to function

   hm  6. jan 2008     rev 1.2
       improved performance

   hm  26. oct. 2008   rev 1.3
       optimized code

   hm  3. nov. 2008    rev 1.4
       used wrong factor in formula

   *)
END_FUNCTION

FUNCTION "SCALE_B8" : Real   // FC333, SCL
TITLE = SCALE_B8
{ S7_Optimized_Access := 'FALSE' }
AUTHOR : hugo
FAMILY : SIGPRO
NAME : SCALEB8
VERSION : 1.4
// this functiob block can scale up to 8 inputs.
// the inputs have their min value at 0 and their max value at 255 while the min and max value can be either positive or negative.
// the inputs ramp between min and max values for the respective inputs to be between (0..255).
// the summed output is then scaled by an scale input K and a offset O can be added to the output.
// the min and max input configurations can be edited in the cfc editor by double clicking the symbol body.
   VAR_INPUT
      in1 : Byte;
      in2 : Byte;
      in3 : Byte;
      in4 : Byte;
      in5 : Byte;
      in6 : Byte;
      in7 : Byte;
      in8 : Byte;
      K : Real;
      O : Real;
      in1_min : Real;
      in1_max : Real;
      in2_min : Real;
      in2_max : Real;
      in3_min : Real;
      in3_max : Real;
      in4_min : Real;
      in4_max : Real;
      in5_min : Real;
      in5_max : Real;
      in6_min : Real;
      in6_max : Real;
      in7_min : Real;
      in7_max : Real;
      in8_min : Real;
      in8_max : Real;
   END_VAR
BEGIN


   #SCALE_B8 :=  (((#in1_max - #in1_min)* INT_TO_REAL(BYTE_TO_INT(#in1)) + 
                  (#in2_max - #in2_min)* INT_TO_REAL(BYTE_TO_INT(#in2)) + 
                  (#in3_max - #in3_min)* INT_TO_REAL(BYTE_TO_INT(#in3)) + 
                  (#in4_max - #in4_min)* INT_TO_REAL(BYTE_TO_INT(#in4)) +
                  (#in5_max - #in5_min)* INT_TO_REAL(BYTE_TO_INT(#in5)) + 
                  (#in6_max - #in6_min)* INT_TO_REAL(BYTE_TO_INT(#in6)) + 
                  (#in7_max - #in7_min)* INT_TO_REAL(BYTE_TO_INT(#in7)) + 
                  (#in8_max - #in8_min)* INT_TO_REAL(BYTE_TO_INT(#in8))) * 0.003921569 + 
                  #in1_min + #in2_min + #in3_min + #in4_min + #in5_min + #in6_min + #in7_min + #in8_min) * #K + #O;


   (* revision History
   hm  19. jan.2007    rev 1.1
       changed outputs to real to avoid overflow of integer
       added offset for better cascading of scale functions

   hm  6. jan. 2008    rev 1.2
       improved performance

   hm  26. oct. 2008   rev 1.3
       code optimization

   hm  3. nov. 2008    rev 1.4
       used wrong factor in formula

   *)
END_FUNCTION